VERSION : 0.1
   VAR_INPUT
      OFF_SQ : Bool := false;   // Turn sequence off
      INIT_SQ : Bool := false;   // Set sequence to initial state
      ACK_EF : Bool := false;   // Acknowledge all errors and faults
   END_VAR
   VAR_OUTPUT
      S_NO : Int := 0;   // Step number
      S_MORE : Bool := false;   // More steps are available and can be shown in S_NO
      S_ACTIVE : Bool := false;   // Step indicated in S_NO is active
      ERR_FLT : Bool := false;   // Interlock or supervision group error
      AUTO_ON : Bool := false;   // Automatic mode is active
   END_VAR
   VAR
      STATE : Int;   // Step number
      Unit : Struct
         START : Bool;   // Sequence Start
         INITIALIZATION : Bool;   // Sequence initialization
         ABORTING : Bool;   // Sequence about
         WAIT : Bool;   // Wating for Permissive read only
         COMPLETE : Bool;   // Sequence done
         "TURN ON" : Bool;   // Operator turn on retail equiment Button
         "TURN OFF" : Bool;   // Operator turn off retail equiment Button
         DONE : Bool;   // Operator Material is Being remove Button
         LV : Bool;
         PM : Bool;
         OverFlowCheck : Struct   // Check the Centrifuge is not over Material
            Enable : Bool;
            Wait_over : Bool;
            wait_pmp : Bool;
         END_STRUCT;
         TURBIDITY : Struct
            Enable : Bool;
            Wait : Bool;
         END_STRUCT;
         "WET CAKE_DRAIN" : Bool;
         Flow_SP : Real := 5.0;   // L/Min Flow Setpoint for FV-3011
         "TIMER" : Struct
            BucketTimer : IEC_TIMER;
            "WET-CAKE" : IEC_TIMER;
         END_STRUCT;
         "TIME" : Struct
            "WET-CAKE" : Time := T#10M;
            CountDown : Struct
               "WET-CAKE" : Time;
            END_STRUCT;
         END_STRUCT;
      END_STRUCT;
      HMI_INFO : Array[0..11] of UInt;
      IF_PAR : G7_IfParPlus_V6;
      RT_DATA : G7_RTDataPlus_V6;   // Internal data area
      Abort : G7_TransitionPlus_V6;   // Transition structure
      InitializeR : G7_TransitionPlus_V6;   // Transition structure
      CentfgP : G7_TransitionPlus_V6;   // Transition structure
      Re : G7_TransitionPlus_V6;   // Transition structure
      Centrifuge : G7_TransitionPlus_V6;   // Transition structure
      Wash : G7_TransitionPlus_V6;   // Transition structure
      Std : G7_TransitionPlus_V6;   // Transition structure
      StT : G7_TransitionPlus_V6;   // Transition structure
      MotorOn : G7_TransitionPlus_V6;   // Transition structure
      ROpnd : G7_TransitionPlus_V6;   // Transition structure
      AutoFlw : G7_TransitionPlus_V6;   // Transition structure
      TOT_Dn : G7_TransitionPlus_V6;   // Transition structure
      TransfDn : G7_TransitionPlus_V6;   // Transition structure
      TnkIdle : G7_TransitionPlus_V6;   // Transition structure
      WaterDn : G7_TransitionPlus_V6;   // Transition structure
      WtPmOff : G7_TransitionPlus_V6;   // Transition structure
      BcketTDn : G7_TransitionPlus_V6;   // Transition structure
      PmpsOff : G7_TransitionPlus_V6;   // Transition structure
      CntrfgOff : G7_TransitionPlus_V6;   // Transition structure
      CntrfgEnd : G7_TransitionPlus_V6;   // Transition structure
      Init : G7_TransitionPlus_V6;   // Transition structure
      SAut : G7_TransitionPlus_V6;   // Transition structure
      SIn : G7_TransitionPlus_V6;   // Transition structure
      Initd : G7_TransitionPlus_V6;   // Transition structure
      Trans145 : G7_TransitionPlus_V6;   // Transition structure
      Ab : G7_TransitionPlus_V6;   // Transition structure
      AbortOn : G7_TransitionPlus_V6;   // Transition structure
      AbortDn : G7_TransitionPlus_V6;   // Transition structure
      Idle : G7_StepPlus_V6;   // Step structure
      Ready : G7_StepPlus_V6;   // Step structure
      SelectSeq : G7_StepPlus_V6;   // Step structure
      Started : G7_StepPlus_V6;   // Step structure
      StartTank : G7_StepPlus_V6;   // Step structure
      "USER CentrOn" : G7_StepPlus_V6;   // Step structure
      OpenRoute : G7_StepPlus_V6;   // Step structure
      AutoFlowCtl : G7_StepPlus_V6;   // Step structure
      Transfering : G7_StepPlus_V6;   // Step structure
      Complete : G7_StepPlus_V6;   // Step structure
      ReleaseTank : G7_StepPlus_V6;   // Step structure
      "USER SlWash" : G7_StepPlus_V6;   // Step structure
      StopReqWater : G7_StepPlus_V6;   // Step structure
      Drying : G7_StepPlus_V6;   // Step structure
      DryingDone : G7_StepPlus_V6;   // Step structure
      "USER CentrOff" : G7_StepPlus_V6;   // Step structure
      End : G7_StepPlus_V6;   // Step structure
      Initialize : G7_StepPlus_V6;   // Step structure
      SetAuto : G7_StepPlus_V6;   // Step structure
      SetInitial : G7_StepPlus_V6;   // Step structure
      "2ndReset" : G7_StepPlus_V6;   // Step structure
      FeelerEngage : G7_StepPlus_V6;   // Step structure
      AbortStarting : G7_StepPlus_V6;   // Step structure
      Aborting : G7_StepPlus_V6;   // Step structure
      AbortDone : G7_StepPlus_V6;   // Step structure
      SINI : Array[0..4] of USInt;
      LSTT : Array[0..27] of USInt;
      ATAJ : Array[0..27] of USInt;
      ATAB : Array[0..27] of USInt;
      PSTT : Array[0..27] of USInt;
      NSTT : Array[0..27] of USInt;
      ASSJ : Array[0..24] of USInt;
      ASSB : Array[0..24] of USInt;
      PTTS : Array[0..24] of USInt;
      NTTS : Array[0..24] of USInt;
      SW_SQTS : Array[0..24] of USInt;
      SWITCH : Array[0..3] of USInt;
      TVX : Array[0..9] of USInt;
      TTX : Array[0..9] of USInt;
      TSX : Array[0..4] of USInt;
      S00X : Array[0..4] of USInt;
      SOFFX : Array[0..4] of USInt;
      SONX : Array[0..4] of USInt;
      SAX : Array[0..4] of USInt;
      SERRX : Array[0..25] of USInt;
      SMX : Array[0..25] of USInt;
      S0X : Array[0..25] of USInt;
      S1X : Array[0..25] of USInt;
      IL_ALARM_INST : Diag_Alarm;
      SUP_ALARM_INST : Diag_Alarm;
      STEP_TIME_ALARM_INST : Diag_Alarm;
      IEC_TIMER_INST : IEC_TIMER;
      TRANSACTION_FLAG : Bool := false;
   END_VAR
   // LSTT[8] := 255;
   // SINI[0] := 2;
   // LSTT[0] := 22;
   // NSTT[0] := 22;
   // PTTS[0] := 255;
   // TVX[0] := 16#1;
   // TTX[0] := 16#1;
   // TSX[0] := 16#1;
   // S00X[0] := 16#1;
   // SOFFX[0] := 16#1;
   // SONX[0] := 16#1;
   // SAX[0] := 16#1;
   // SERRX[0] := 16#1;
   // SMX[0] := 16#1;
   // S0X[0] := 16#1;
   // S1X[0] := 16#1;
   // LSTT[1] := 17;
   // LSTT[2] := 255;
   // LSTT[3] := 255;
   // LSTT[4] := 3;
   // LSTT[5] := 255;
   // LSTT[6] := 255;
   // LSTT[7] := 255;
   // LSTT[9] := 255;
   // LSTT[13] := 255;
   // LSTT[10] := 255;
   // LSTT[11] := 255;
   // LSTT[12] := 255;
   // NSTT[8] := 6;
   // LSTT[14] := 255;
   // LSTT[15] := 255;
   // LSTT[16] := 255;
   // LSTT[17] := 255;
   // LSTT[18] := 255;
   // ATAJ[1] := 1;
   // ATAJ[2] := 2;
   // ATAJ[3] := 3;
   // ATAJ[4] := 4;
   // ATAJ[5] := 5;
   // ATAJ[6] := 6;
   // ATAJ[7] := 7;
   // ATAJ[8] := 8;
   // ATAJ[9] := 9;
   // ATAJ[10] := 10;
   // ATAJ[11] := 11;
   // ATAJ[12] := 12;
   // ATAJ[13] := 13;
   // ATAJ[14] := 14;
   // ATAJ[15] := 15;
   // ATAJ[16] := 16;
   // ATAJ[17] := 17;
   // ATAJ[18] := 18;
   // ATAJ[19] := 19;
   // ATAB[1] := 2;
   // ATAB[17] := 17;
   // ATAB[3] := 3;
   // ATAB[4] := 5;
   // ATAB[5] := 4;
   // ATAB[6] := 6;
   // ATAB[7] := 7;
   // ATAB[8] := 8;
   // ATAB[9] := 9;
   // ATAB[10] := 10;
   // ATAB[11] := 11;
   // ATAB[12] := 12;
   // ATAB[13] := 13;
   // ATAB[14] := 14;
   // ATAB[15] := 15;
   // ATAB[16] := 16;
   // ATAB[19] := 19;
   // ATAB[18] := 18;
   // PSTT[17] := 14;
   // PSTT[14] := 11;
   // PSTT[3] := 1;
   // PSTT[4] := 2;
   // PSTT[5] := 2;
   // PSTT[6] := 3;
   // PSTT[7] := 4;
   // PSTT[8] := 5;
   // PSTT[9] := 6;
   // PSTT[10] := 7;
   // PSTT[11] := 8;
   // PSTT[12] := 9;
   // PSTT[13] := 10;
   // PSTT[15] := 12;
   // PSTT[16] := 13;
   // PSTT[19] := 16;
   // PSTT[18] := 15;
   // PSTT[21] := 18;
   // NSTT[1] := 17;
   // NSTT[2] := 1;
   // NSTT[3] := 2;
   // NSTT[4] := 3;
   // NSTT[5] := 255;
   // NSTT[6] := 4;
   // NSTT[7] := 5;
   // NSTT[9] := 7;
   // NSTT[13] := 11;
   // NSTT[10] := 8;
   // NSTT[11] := 9;
   // NSTT[12] := 10;
   // NSTT[14] := 12;
   // NSTT[15] := 13;
   // NSTT[16] := 14;
   // NSTT[17] := 15;
   // NSTT[18] := 16;
   // ASSJ[1] := 1;
   // ASSJ[2] := 2;
   // ASSJ[3] := 3;
   // ASSJ[4] := 4;
   // ASSJ[5] := 5;
   // ASSJ[6] := 6;
   // ASSJ[7] := 7;
   // ASSJ[8] := 8;
   // ASSJ[9] := 9;
   // ASSJ[10] := 10;
   // ASSJ[11] := 11;
   // ASSJ[12] := 12;
   // ASSJ[13] := 13;
   // ASSJ[14] := 14;
   // ASSJ[15] := 15;
   // ASSJ[16] := 16;
   // ASSB[1] := 1;
   // ASSB[2] := 2;
   // ASSB[3] := 3;
   // ASSB[4] := 4;
   // ASSB[5] := 5;
   // ASSB[6] := 6;
   // ASSB[7] := 7;
   // ASSB[8] := 8;
   // ASSB[9] := 9;
   // ASSB[10] := 10;
   // ASSB[11] := 11;
   // ASSB[12] := 12;
   // ASSB[13] := 13;
   // ASSB[14] := 14;
   // ASSB[15] := 15;
   // ASSB[16] := 16;
   // PTTS[2] := 3;
   // PTTS[3] := 255;
   // PTTS[4] := 6;
   // PTTS[5] := 7;
   // PTTS[6] := 8;
   // PTTS[7] := 9;
   // PTTS[8] := 10;
   // PTTS[9] := 11;
   // PTTS[10] := 12;
   // PTTS[11] := 13;
   // PTTS[12] := 14;
   // PTTS[13] := 15;
   // PTTS[14] := 16;
   // PTTS[15] := 17;
   // PTTS[16] := 18;
   // NTTS[1] := 3;
   // NTTS[2] := 4;
   // NTTS[3] := 6;
   // NTTS[4] := 7;
   // NTTS[5] := 8;
   // NTTS[6] := 9;
   // NTTS[7] := 10;
   // NTTS[8] := 11;
   // NTTS[9] := 12;
   // NTTS[10] := 13;
   // NTTS[11] := 14;
   // NTTS[12] := 15;
   // NTTS[13] := 16;
   // NTTS[14] := 17;
   // NTTS[15] := 18;
   // NTTS[16] := 19;
   // SW_SQTS[6] := 2;
   // SW_SQTS[7] := 2;
   // SW_SQTS[8] := 2;
   // SW_SQTS[9] := 2;
   // SW_SQTS[10] := 2;
   // SW_SQTS[11] := 2;
   // SW_SQTS[12] := 2;
   // SW_SQTS[13] := 2;
   // SW_SQTS[14] := 2;
   // SW_SQTS[15] := 2;
   // SW_SQTS[16] := 2;
   // NTTS[23] := 26;
   // NTTS[22] := 25;
   // NTTS[21] := 24;
   // NTTS[20] := 23;
   // NTTS[19] := 22;
   // NTTS[18] := 21;
   // NTTS[17] := 20;
   // PTTS[23] := 25;
   // PTTS[22] := 255;
   // PTTS[21] := 23;
   // PTTS[20] := 22;
   // PTTS[19] := 21;
   // PTTS[18] := 20;
   // PTTS[17] := 255;
   // ASSB[23] := 23;
   // ASSB[22] := 22;
   // ASSB[21] := 21;
   // ASSB[20] := 20;
   // ASSB[19] := 19;
   // ASSB[18] := 18;
   // ASSB[17] := 17;
   // ASSJ[23] := 23;
   // ASSJ[22] := 22;
   // ASSJ[21] := 21;
   // ASSJ[20] := 20;
   // ASSJ[19] := 19;
   // ASSJ[18] := 18;
   // ASSJ[17] := 17;
   // NSTT[23] := 21;
   // NSTT[25] := 23;
   // PSTT[26] := 23;
   // PSTT[25] := 22;
   // PSTT[24] := 21;
   // PSTT[23] := 20;
   // PSTT[22] := 19;
   // PSTT[20] := 17;
   // ATAB[26] := 26;
   // ATAB[25] := 25;
   // ATAB[24] := 24;
   // ATAB[23] := 23;
   // ATAB[22] := 22;
   // ATAB[21] := 21;
   // ATAB[20] := 20;
   // ATAJ[26] := 26;
   // ATAJ[25] := 25;
   // ATAJ[24] := 24;
   // ATAJ[23] := 23;
   // ATAJ[22] := 22;
   // ATAJ[21] := 21;
   // ATAJ[20] := 20;
   // LSTT[23] := 255;
   // LSTT[25] := 255;
   // SW_SQTS[17] := 3;
   // SW_SQTS[18] := 3;
   // SW_SQTS[19] := 3;
   // SW_SQTS[20] := 3;
   // SW_SQTS[21] := 3;
   // SW_SQTS[22] := 4;
   // SW_SQTS[23] := 4;
   // SINI[2] := 255;
   // SINI[3] := 255;
   // LSTT[21] := 255;
   // NSTT[21] := 19;
   // SW_SQTS[2] := 1;
   // SW_SQTS[3] := 2;
   // SW_SQTS[4] := 2;
   // SW_SQTS[5] := 2;
   // Unit."TIMER".BucketTimer.PT := T#10S;
   // LSTT[24] := 1;
   // LSTT[22] := 255;
   // NSTT[22] := 20;
   // NSTT[24] := 1;
   // Unit."TIMER"."WET-CAKE".PT := T#10M;
   // SINI[4] := 255;
   // LSTT[20] := 255;
   // NSTT[20] := 18;
   // PTTS[1] := 2;
   // SWITCH[1] := 239;
   // SWITCH[0] := 156;
   // SWITCH[2] := 251;
   // ATAB[0] := 1;
   // SW_SQTS[1] := 1;
   // LSTT[26] := 255;
   // ATAJ[27] := 27;
   // ATAB[27] := 27;
   // PSTT[27] := 24;
   // NSTT[26] := 24;
   // ASSJ[24] := 24;
   // ASSB[24] := 24;
   // PTTS[24] := 26;
   // NTTS[24] := 27;
   // SW_SQTS[24] := 4;
BEGIN
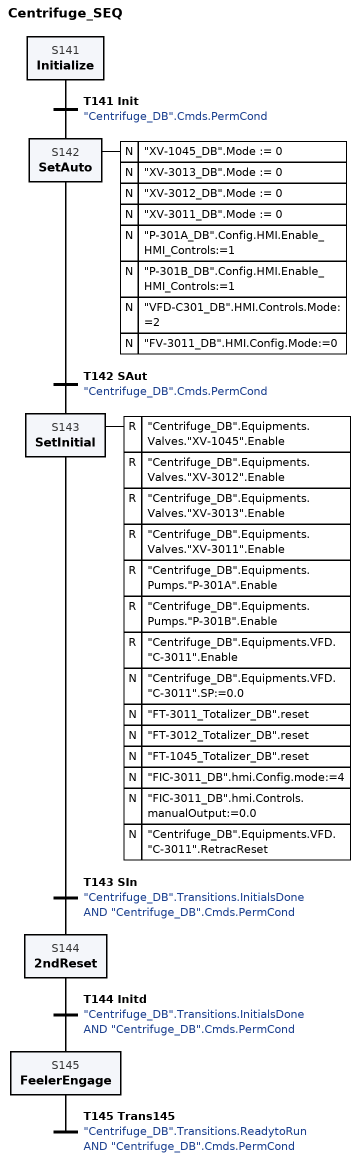
   // permanent pre-instructions
   NETWORK 1
      "Centrifuge_Signals_FROM_T-103"();
      "Centrifuge_Signals_FROM_T-104"();
      "Centrifuge_SEQ_FC"();
      "Centrifuge_Transitions_FC"();

   // sequencer 1
   STEP "2ndReset":   // S144, max time T#10S, warning time T#7S
      // Initialize T-101 Batch sequence
   END_STEP
   TRANSITION Initd FROM "2ndReset" TO FeelerEngage   // T144
      := "Centrifuge_DB".Transitions.InitialsDone AND "Centrifuge_DB".Cmds.PermCond;
   END_TRANSITION
   STEP Initialize:   // S141, max time T#10S, warning time T#7S
      // Initialize T-101 Batch sequence
   END_STEP
   TRANSITION Init FROM Initialize TO SetAuto   // T141: CLOSED: XV-1041
      := "Centrifuge_DB".Cmds.PermCond;
   END_TRANSITION
   STEP SetInitial:   // S143, max time T#10S, warning time T#7S
      // Initialize T-101 Batch sequence
              R    "Centrifuge_DB".Equipments.Valves."XV-1045".Enable
              R    "Centrifuge_DB".Equipments.Valves."XV-3012".Enable
              R    "Centrifuge_DB".Equipments.Valves."XV-3013".Enable
              R    "Centrifuge_DB".Equipments.Valves."XV-3011".Enable
              R    "Centrifuge_DB".Equipments.Pumps."P-301A".Enable
              R    "Centrifuge_DB".Equipments.Pumps."P-301B".Enable
              R    "Centrifuge_DB".Equipments.VFD."C-3011".Enable
              N    "Centrifuge_DB".Equipments.VFD."C-3011".SP:=0.0
              N    "FT-3011_Totalizer_DB".reset
              N    "FT-3012_Totalizer_DB".reset
              N    "FT-1045_Totalizer_DB".reset
              N    "FIC-3011_DB".hmi.Config.mode:=4
              N    "FIC-3011_DB".hmi.Controls.manualOutput:=0.0
              N    "Centrifuge_DB".Equipments.VFD."C-3011".RetracReset
   END_STEP
   TRANSITION SIn FROM SetInitial TO "2ndReset"   // T143: CLOSED: XV-1013
      := "Centrifuge_DB".Transitions.InitialsDone AND "Centrifuge_DB".Cmds.PermCond;
   END_TRANSITION
   STEP SetAuto:   // S142, max time T#10S, warning time T#7S
              N    "XV-1045_DB".Mode := 0
              N    "XV-3013_DB".Mode := 0
              N    "XV-3012_DB".Mode := 0
              N    "XV-3011_DB".Mode := 0
              N    "P-301A_DB".Config.HMI.Enable_HMI_Controls:=1
              N    "P-301B_DB".Config.HMI.Enable_HMI_Controls:=1
              N    "VFD-C301_DB".HMI.Controls.Mode:=2
              N    "FV-3011_DB".HMI.Config.Mode:=0
   END_STEP
   TRANSITION SAut FROM SetAuto TO SetInitial   // T142
      := "Centrifuge_DB".Cmds.PermCond;
   END_TRANSITION
   STEP FeelerEngage:   // S145, max time T#10S, warning time T#7S
   END_STEP
   TRANSITION Trans145 FROM FeelerEngage TO ?   // T145
      := "Centrifuge_DB".Transitions.ReadytoRun AND "Centrifuge_DB".Cmds.PermCond;
   END_TRANSITION

   // permanent post-instructions
   NETWORK 1
      "Centrifuge_FC_Outputs"();
END_FUNCTION_BLOCK

FUNCTION "Centrifuge_SEQ_FC_old" : Void   // FC75, LAD
{ S7_Optimized_Access := 'TRUE' }
VERSION : 0.1
   VAR_TEMP   // added for the SCL form of the ladder/FBD networks
      _w1 : Bool;
      _w2 : Bool;
   END_VAR
BEGIN

REGION Network 2: Abort
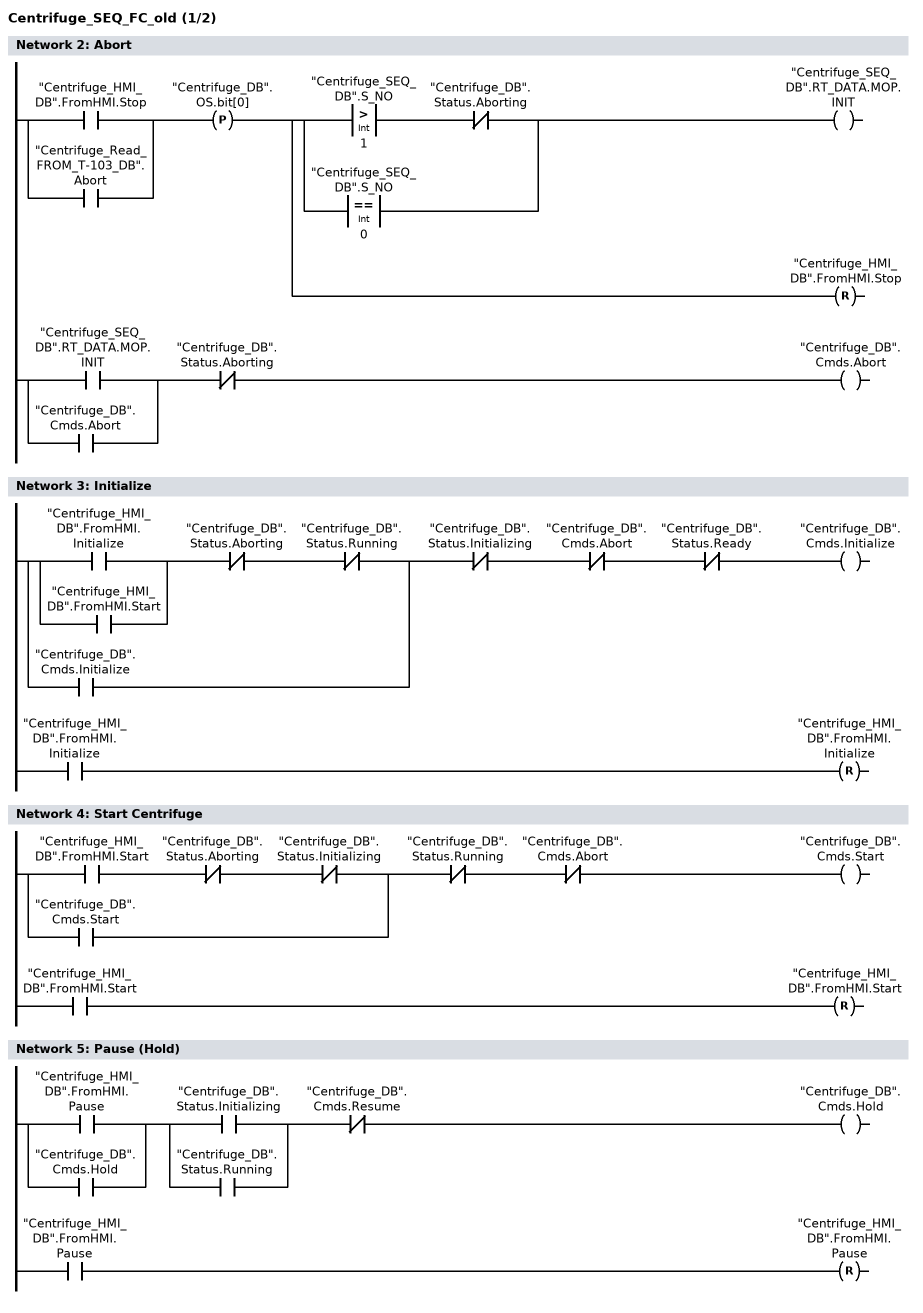
   RUNG wire#powerrail
      Contact( "Centrifuge_HMI_DB".FromHMI.Stop )
      wire#w1
      P_Trig( "Centrifuge_DB".OS.bit[0] )
      wire#w2
      { S7_Templates := "SrcType := Int" } GT_Contact(in1 := "Centrifuge_SEQ_DB".S_NO, in2 := 1)
      I_Contact( "Centrifuge_DB".Status.Aborting )
      wire#w3
      Coil( "Centrifuge_SEQ_DB".RT_DATA.MOP.INIT )
   END_RUNG
   RUNG wire#powerrail
      Contact( "Centrifuge_Read_FROM_T-103_DB".Abort )
   END_RUNG wire#w1
   RUNG wire#w2
      { S7_Templates := "SrcType := Int" } EQ_Contact(in1 := "Centrifuge_SEQ_DB".S_NO, in2 := 0)
   END_RUNG wire#w3
   RUNG wire#w2
      R_Coil( "Centrifuge_HMI_DB".FromHMI.Stop )
   END_RUNG
   RUNG wire#powerrail
      Contact( "Centrifuge_SEQ_DB".RT_DATA.MOP.INIT )
      wire#w4
      I_Contact( "Centrifuge_DB".Status.Aborting )
      Coil( "Centrifuge_DB".Cmds.Abort )
   END_RUNG
   RUNG wire#powerrail
      Contact( "Centrifuge_DB".Cmds.Abort )
   END_RUNG wire#w4
   // the same network as SCL:
   #_w1 := "Centrifuge_HMI_DB".FromHMI.Stop OR "Centrifuge_Read_FROM_T-103_DB".Abort;
   #_w2 := #_w1 AND NOT "Centrifuge_DB".OS.bit[0];   // rising edge
   "Centrifuge_DB".OS.bit[0] := #_w1;
   "Centrifuge_SEQ_DB".RT_DATA.MOP.INIT := #_w2 AND ((("Centrifuge_SEQ_DB".S_NO > 1) AND NOT "Centrifuge_DB".Status.Aborting) OR ("Centrifuge_SEQ_DB".S_NO = 0));
   IF #_w2 THEN "Centrifuge_HMI_DB".FromHMI.Stop := FALSE; END_IF;
   "Centrifuge_DB".Cmds.Abort := ("Centrifuge_SEQ_DB".RT_DATA.MOP.INIT OR "Centrifuge_DB".Cmds.Abort) AND NOT "Centrifuge_DB".Status.Aborting;
END_REGION

REGION Network 3: Initialize
   RUNG wire#powerrail
      Contact( "Centrifuge_HMI_DB".FromHMI.Initialize )
      wire#w1
      I_Contact( "Centrifuge_DB".Status.Aborting )
      I_Contact( "Centrifuge_DB".Status.Running )
      wire#w2
      I_Contact( "Centrifuge_DB".Status.Initializing )
      I_Contact( "Centrifuge_DB".Cmds.Abort )
      I_Contact( "Centrifuge_DB".Status.Ready )
      Coil( "Centrifuge_DB".Cmds.Initialize )
   END_RUNG
   RUNG wire#powerrail
      Contact( "Centrifuge_HMI_DB".FromHMI.Start )
   END_RUNG wire#w1
   RUNG wire#powerrail
      Contact( "Centrifuge_DB".Cmds.Initialize )
   END_RUNG wire#w2
   RUNG wire#powerrail
      Contact( "Centrifuge_HMI_DB".FromHMI.Initialize )
      R_Coil( "Centrifuge_HMI_DB".FromHMI.Initialize )
   END_RUNG
   // the same network as SCL:
   "Centrifuge_DB".Cmds.Initialize := ((("Centrifuge_HMI_DB".FromHMI.Initialize OR "Centrifuge_HMI_DB".FromHMI.Start) AND NOT "Centrifuge_DB".Status.Aborting AND NOT "Centrifuge_DB".Status.Running) OR "Centrifuge_DB".Cmds.Initialize) AND NOT "Centrifuge_DB".Status.Initializing AND NOT "Centrifuge_DB".Cmds.Abort AND NOT "Centrifuge_DB".Status.Ready;
   IF "Centrifuge_HMI_DB".FromHMI.Initialize THEN "Centrifuge_HMI_DB".FromHMI.Initialize := FALSE; END_IF;
END_REGION

REGION Network 4: Start Centrifuge
   RUNG wire#powerrail
      Contact( "Centrifuge_HMI_DB".FromHMI.Start )
      I_Contact( "Centrifuge_DB".Status.Aborting )
      I_Contact( "Centrifuge_DB".Status.Initializing )
      wire#w1
      I_Contact( "Centrifuge_DB".Status.Running )
      I_Contact( "Centrifuge_DB".Cmds.Abort )
      Coil( "Centrifuge_DB".Cmds.Start )
   END_RUNG
   RUNG wire#powerrail
      Contact( "Centrifuge_DB".Cmds.Start )
   END_RUNG wire#w1
   RUNG wire#powerrail
      Contact( "Centrifuge_HMI_DB".FromHMI.Start )
      R_Coil( "Centrifuge_HMI_DB".FromHMI.Start )
   END_RUNG
   // the same network as SCL:
   "Centrifuge_DB".Cmds.Start := (("Centrifuge_HMI_DB".FromHMI.Start AND NOT "Centrifuge_DB".Status.Aborting AND NOT "Centrifuge_DB".Status.Initializing) OR "Centrifuge_DB".Cmds.Start) AND NOT "Centrifuge_DB".Status.Running AND NOT "Centrifuge_DB".Cmds.Abort;
   IF "Centrifuge_HMI_DB".FromHMI.Start THEN "Centrifuge_HMI_DB".FromHMI.Start := FALSE; END_IF;
END_REGION

REGION Network 5: Pause (Hold)
   RUNG wire#powerrail
      Contact( "Centrifuge_HMI_DB".FromHMI.Pause )
      wire#w1
      Contact( "Centrifuge_DB".Status.Initializing )
      wire#w2
      I_Contact( "Centrifuge_DB".Cmds.Resume )
      Coil( "Centrifuge_DB".Cmds.Hold )
   END_RUNG
   RUNG wire#powerrail
      Contact( "Centrifuge_DB".Cmds.Hold )
   END_RUNG wire#w1
   RUNG wire#w1
      Contact( "Centrifuge_DB".Status.Running )
   END_RUNG wire#w2
   RUNG wire#powerrail
      Contact( "Centrifuge_HMI_DB".FromHMI.Pause )
      R_Coil( "Centrifuge_HMI_DB".FromHMI.Pause )
   END_RUNG
   // the same network as SCL:
   "Centrifuge_DB".Cmds.Hold := ("Centrifuge_HMI_DB".FromHMI.Pause OR "Centrifuge_DB".Cmds.Hold) AND ("Centrifuge_DB".Status.Initializing OR "Centrifuge_DB".Status.Running) AND NOT "Centrifuge_DB".Cmds.Resume;
   IF "Centrifuge_HMI_DB".FromHMI.Pause THEN "Centrifuge_HMI_DB".FromHMI.Pause := FALSE; END_IF;
END_REGION

REGION Network 6: Restart From Pause (Hold)
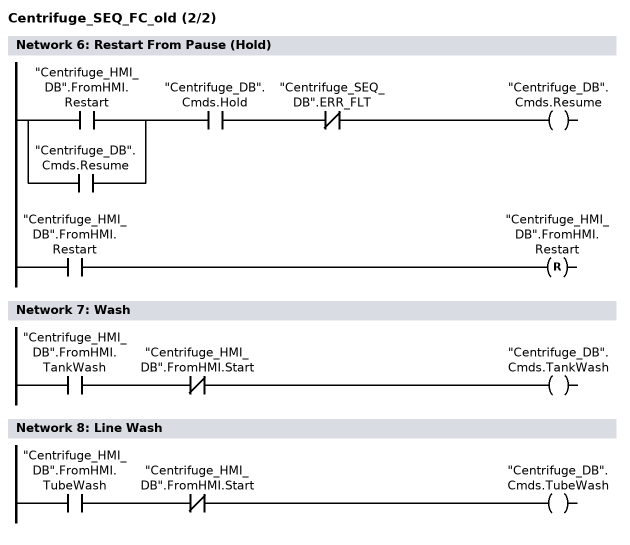
   RUNG wire#powerrail
      Contact( "Centrifuge_HMI_DB".FromHMI.Restart )
      wire#w1
      Contact( "Centrifuge_DB".Cmds.Hold )
      I_Contact( "Centrifuge_SEQ_DB".ERR_FLT )
      Coil( "Centrifuge_DB".Cmds.Resume )
   END_RUNG
   RUNG wire#powerrail
      Contact( "Centrifuge_DB".Cmds.Resume )
   END_RUNG wire#w1
   RUNG wire#powerrail
      Contact( "Centrifuge_HMI_DB".FromHMI.Restart )
      R_Coil( "Centrifuge_HMI_DB".FromHMI.Restart )
   END_RUNG
   // the same network as SCL:
   "Centrifuge_DB".Cmds.Resume := ("Centrifuge_HMI_DB".FromHMI.Restart OR "Centrifuge_DB".Cmds.Resume) AND "Centrifuge_DB".Cmds.Hold AND NOT "Centrifuge_SEQ_DB".ERR_FLT;
   IF "Centrifuge_HMI_DB".FromHMI.Restart THEN "Centrifuge_HMI_DB".FromHMI.Restart := FALSE; END_IF;
END_REGION

REGION Network 7: Wash
   RUNG wire#powerrail
      Contact( "Centrifuge_HMI_DB".FromHMI.TankWash )
      I_Contact( "Centrifuge_HMI_DB".FromHMI.Start )
      Coil( "Centrifuge_DB".Cmds.TankWash )
   END_RUNG
   // the same network as SCL:
   "Centrifuge_DB".Cmds.TankWash := "Centrifuge_HMI_DB".FromHMI.TankWash AND NOT "Centrifuge_HMI_DB".FromHMI.Start;
END_REGION

REGION Network 8: Line Wash
   RUNG wire#powerrail
      Contact( "Centrifuge_HMI_DB".FromHMI.TubeWash )
      I_Contact( "Centrifuge_HMI_DB".FromHMI.Start )
      Coil( "Centrifuge_DB".Cmds.TubeWash )
   END_RUNG
   // the same network as SCL:
   "Centrifuge_DB".Cmds.TubeWash := "Centrifuge_HMI_DB".FromHMI.TubeWash AND NOT "Centrifuge_HMI_DB".FromHMI.Start;
END_REGION

REGION Network 9 (SCL): Sequence Status
   IF "Centrifuge_SEQ_DB".S_NO= 1 THEN
       "Centrifuge_DB".Status.Status := 1; //Idle
   ELSIF "Centrifuge_SEQ_DB".S_NO > 1 AND "Centrifuge_SEQ_DB".S_NO < 150 AND NOT "Centrifuge_SEQ_DB".ERR_FLT THEN
       "Centrifuge_DB".Status.Status := 2; //Running
   ELSIF "Centrifuge_SEQ_DB".S_NO >= 151 AND "Centrifuge_SEQ_DB".S_NO <= 160 AND NOT "Centrifuge_SEQ_DB".ERR_FLT THEN
       "Centrifuge_DB".Status.Status := 3; // Stopping
   ELSIF ("Centrifuge_SEQ_DB".ERR_FLT OR "Centrifuge_DB".Cmds.Hold)  AND "Centrifuge_DB".Status.Status =2 THEN
       "Centrifuge_DB".Status.Status := 4; //Held
   ELSIF ("Centrifuge_SEQ_DB".ERR_FLT OR "Centrifuge_DB".Cmds.Hold) AND  "Centrifuge_DB".Status.Status =2 AND "Centrifuge_Aux_DB"."Bool".TOff  THEN
       "Centrifuge_DB".Status.Status := 5; // Holding
   ELSE
       "Centrifuge_DB".Status.Status := 6; //Unknown
   END_IF;

   //Enable/Disable HMI Start/Stop Button
   "Centrifuge_HMI_DB".ToHMI.EnStopButton := ("Centrifuge_DB".Status.Status > 1) OR "Centrifuge_DB".Status.Step = 0; //Enable HMI Stop Button
   "Centrifuge_HMI_DB".ToHMI.EnStartButton := "Centrifuge_DB".Status.Status = 1;   //Enable Start Button
   "Centrifuge_HMI_DB".ToHMI.EnPauseButton := "Centrifuge_DB".Status.Status = 2 AND NOT "Centrifuge_DB".Cmds.Hold; //Enable Pause Button
   "Centrifuge_HMI_DB".ToHMI.EnRestartButton := "Centrifuge_DB".Status.Status = 2 AND "Centrifuge_DB".Cmds.Hold; //Enable Restart Button
END_REGION

REGION Network 10 (SCL): Sequence Step
   "Centrifuge_DB".Status.Step := "Centrifuge_SEQ_DB".S_NO;
END_REGION

REGION Network 11 (SCL): Sequence state (Procedure running)
   IF "Centrifuge_SEQ_DB".S_NO = 3 OR "Centrifuge_SEQ_DB".S_NO = 4 THEN
       "Centrifuge_DB".Status.State := 1; //Ready
   ELSIF "Centrifuge_SEQ_DB".S_NO >= 21 AND "Centrifuge_SEQ_DB".S_NO <= 60 THEN
       "Centrifuge_DB".Status.State := 2; //Mixing 
   ELSIF "Centrifuge_SEQ_DB".S_NO >= 61 AND "Centrifuge_SEQ_DB".S_NO <= 80 THEN
       "Centrifuge_DB".Status.State := 3; //Pouring
   ELSIF "Centrifuge_SEQ_DB".S_NO >= 141 AND "Centrifuge_SEQ_DB".S_NO <= 150 THEN
       "Centrifuge_DB".Status.State := 4; //Initializing
   ELSIF "Centrifuge_SEQ_DB".S_NO >= 151 AND "Centrifuge_SEQ_DB".S_NO <= 160 THEN
       "Centrifuge_DB".Status.State := 5; //Aborting
   ELSE
       "Centrifuge_DB".Status.State := 0;
   END_IF;
END_REGION

REGION Network 12: Sequence State
END_REGION
END_FUNCTION

FUNCTION "Centrifuge_FC_Outputs" : Void   // FC84, SCL
{ S7_Optimized_Access := 'TRUE' }
VERSION : 0.1
   VAR_TEMP
      Pump_A : Struct
         Cond_01 : Bool;   // Condition 01
         Cond_02 : Bool;
         Cond_03 : Bool;
         Cond_04 : Bool;
      END_STRUCT;
      Pump_B : Struct
         Cond_01 : Bool;   // Condition 01
         Cond_02 : Bool;   // Condition 02
         Cond_03 : Bool;
         Cond_04 : Bool;
         Cond_05 : Bool;
      END_STRUCT;
      Motor : Struct
         Cond_01 : Bool;   // Condition 01
         Cond_02 : Bool;   // Condition 02
      END_STRUCT;
      XV : Struct
         "1045" : Bool;
         "3011" : Bool;
         "3012" : Bool;
         "3013" : Bool;
      END_STRUCT;
      "FV-3011" : Struct
         On : Bool;
         Cond_1 : Bool;
      END_STRUCT;
   END_VAR
BEGIN
   //****** Equipmens Activation*******
   //
   //**************************************************************
   //

   //IF "AlwaysFALSE"  AND  ("Centrifuge_DB".Status.Status <> 1) THEN

       //***********************************************Water Inlet Valve**********************************************************************
       IF "XV-1045_DB".Mode = 0 THEN
           "Centrifuge_DB".Equipments.Valves."XV-1045".CmdOn := "Centrifuge_DB".Equipments.Valves."XV-1045".Enable 
           AND "ZT-C301_DB".SAI>"CentrifugeSpeed" AND NOT "Centrifuge_DB".Cmds.Hold;
           //Delay Off To avoid Overpressure the Lines
           #XV."1045" := "Centrifuge_DB".Equipments.Valves."XV-1045".CmdOn;
           "Centrifuge_Aux_DB".Timer."XV-1045".TOF(IN := #XV."1045",
                                                   PT := "Centrifuge_Aux_DB".Constants.CmdDelay);
           //Command to the Valve
           IF "Centrifuge_Aux_DB".Timer."XV-1045".Q THEN
               "XV-1045_DB".CMD := 2;
           ELSE
               "XV-1045_DB".CMD := 1;
           END_IF;
           "Centrifuge_DB".Equipments.Valves."XV-1045".TurningOff := NOT "Centrifuge_DB".Equipments.Valves."XV-1045".CmdOn AND "Centrifuge_Aux_DB".Timer."XV-1045".Q;
       END_IF;
       //***********************************************Inlet Valve**********************************************************************
       IF "XV-3011_DB".Mode = 0 THEN
           "Centrifuge_DB".Equipments.Valves."XV-3011".CmdOn := "Centrifuge_DB".Equipments.Valves."XV-3011".Enable
           AND NOT "Centrifuge_Aux_DB"."Bool".Centrifuge.Status.FeelerRetracted  AND NOT "Centrifuge_DB".Cmds.Hold;
           //Delay Off To avoid Overpressure the Lines
           #XV."3011" := "Centrifuge_DB".Equipments.Valves."XV-3011".CmdOn;
           "Centrifuge_Aux_DB".Timer."XV-3011".TOF(IN := #XV."3011",
           PT := "Centrifuge_Aux_DB".Constants.CmdDelay);
           IF "Centrifuge_Aux_DB".Timer."XV-3011".Q THEN
               "XV-3011_DB".CMD := 2;
           ELSE
               "XV-3011_DB".CMD := 1;
           END_IF;
           "Centrifuge_DB".Equipments.Valves."XV-3011".TurningOff := NOT "Centrifuge_DB".Equipments.Valves."XV-3011".CmdOn AND "Centrifuge_Aux_DB".Timer."XV-3011".Q;
       END_IF;
       //***********************************************Return Valve**********************************************************************
       IF "XV-3012_DB".Mode = 0 THEN
           "Centrifuge_DB".Equipments.Valves."XV-3012".CmdOn := "Centrifuge_DB".Equipments.Valves."XV-3012".Enable AND NOT "Centrifuge_DB".Cmds.Hold;
           //Delay Off To avoid Overpressure the Lines
           #XV."3012" := "Centrifuge_DB".Equipments.Valves."XV-3012".CmdOn;
           "Centrifuge_Aux_DB".Timer."XV-3012".TOF(IN := #XV."3012",
                                                   PT := "Centrifuge_Aux_DB".Constants.CmdDelay);
           //Command to the Valve
           IF "Centrifuge_Aux_DB".Timer."XV-3012".Q THEN
               "XV-3012_DB".CMD := 2;
           ELSE
               "XV-3012_DB".CMD := 1;
           END_IF;
           "Centrifuge_DB".Equipments.Valves."XV-3012".TurningOff := NOT "Centrifuge_DB".Equipments.Valves."XV-3012".CmdOn AND "Centrifuge_Aux_DB".Timer."XV-3012".Q;
       END_IF;
       //***********************************************Outlet Valve**********************************************************************
       IF "XV-3013_DB".Mode = 0 THEN
           "Centrifuge_DB".Equipments.Valves."XV-3013".CmdOn := "Centrifuge_DB".Equipments.Valves."XV-3013".Enable AND NOT "Centrifuge_DB".Cmds.Hold;
           //Delay Off To avoid Overpressure the Lines
           #XV."3013" := "Centrifuge_DB".Equipments.Valves."XV-3013".CmdOn;
           "Centrifuge_Aux_DB".Timer."XV-3013".TOF(IN := #XV."3013",
                                                   PT := "Centrifuge_Aux_DB".Constants.CmdDelay);
           //Command to the Valve
           IF "Centrifuge_Aux_DB".Timer."XV-3013".Q THEN
               "XV-3013_DB".CMD := 2;
           ELSE
               "XV-3013_DB".CMD := 1;
           END_IF;
           "Centrifuge_DB".Equipments.Valves."XV-3013".TurningOff := NOT "Centrifuge_DB".Equipments.Valves."XV-3013".CmdOn AND "Centrifuge_Aux_DB".Timer."XV-3013".Q;
       END_IF;

       //***********************************************FIC-3011 Controller (Centrifuge inlet flow)********************************************************************
       IF "FV-3011_DB".HMI.Config.Mode = 0 THEN
           #"FV-3011".Cond_1 := "Centrifuge_DB".Equipments.Valves."FV-3011".Enable AND "XV-3011_DB".OS;
           "Centrifuge_DB".Equipments.Valves."FV-3011".CmdOn := #"FV-3011".Cond_1 AND NOT "Centrifuge_DB".Cmds.Hold AND NOT "Centrifuge_DB".Status.Aborting;
           //Delay Off To avoid Overpressure the Lines
           #"FV-3011".On := "Centrifuge_DB".Equipments.Valves."FV-3011".CmdOn;
           "Centrifuge_Aux_DB".Timer."FV-3011".TOF(IN := #"FV-3011".On,
                                                   PT := "Centrifuge_Aux_DB".Constants.CmdDelay);
           IF "Centrifuge_Aux_DB".Timer."FV-3011".Q THEN
               "FIC-3011_DB".enableManualMode := False;
               "FIC-3011_DB".enableRemoteSetpoint := False;
               "FIC-3011_DB".hmi.Controls.manualEnable := False;
               "FIC-3011_DB".hmi.Config.mode := 3;
           END_IF;     // ELSE
             //  "FIC-3011_DB".enableManualMode := True;
             //  "FIC-3011_DB".enableRemoteSetpoint := False;
             //  "FIC-3011_DB".hmi.Controls.manualEnable := True;
             //  "FIC-3011_DB".hmi.Config.mode := 4;
            //   "FIC-3011_DB".hmi.Controls.manualOutput := 0;
         //  END_IF;
           "Centrifuge_DB".Equipments.Valves."FV-3011".TurningOff := NOT "Centrifuge_DB".Equipments.Valves."FV-3011".CmdOn AND "Centrifuge_Aux_DB".Timer."FV-3011".Q;
       END_IF;
       // ***********************************************Pump A**********************************************************************
       // Condition to CmdOn "On Command" 
       IF "P-301A_DB".Config.HMI.Enable_HMI_Controls = 1 THEN
           #Pump_A.Cond_01 := "Centrifuge_DB".Equipments.Pumps."P-301A".Enable AND ("Centrifuge_DB".PmpSel."P-301AB" = 1 OR "Centrifuge_DB".PmpSel."P-301AB" = 3);
           #Pump_A.Cond_02 :=  "XV-3013_DB".OS OR "XV-3012_DB".OS; //Outlet Valve Open. 
           #Pump_A.Cond_03 := #Pump_A.Cond_01 AND NOT "Centrifuge_DB".Cmds.Hold;
           "Centrifuge_DB".Equipments.Pumps."P-301A".CmdOn := #Pump_A.Cond_02 AND #Pump_A.Cond_03;
           //**********Commands to the Pumps
           IF "Centrifuge_DB".Equipments.Pumps."P-301A".CmdOn THEN
               "P-301A_DB".Stop_CMD := False;
               "P-301A_DB".Start_CMD := true;
               "P-301A_DB".ON := TRUE;
               "P-301A_DB".OFF := FALSE;
           ELSE
               "P-301A_DB".Stop_CMD := TRUE;
               "P-301A_DB".Start_CMD := FALSE;
               "P-301A_DB".ON := FALSE;
               "P-301A_DB".OFF := TRUE;
           END_IF;
       END_IF;
       // ***********************************************Pump B**********************************************************************
       // Condition to CmdOn "On Command" 
       IF "P-301B_DB".Config.HMI.Enable_HMI_Controls = 1 THEN
           #Pump_B.Cond_01 := "Centrifuge_DB".Equipments.Pumps."P-301B".Enable AND ("Centrifuge_DB".PmpSel."P-301AB" = 2 OR "Centrifuge_DB".PmpSel."P-301AB" = 3);
           #Pump_B.Cond_02 := "XV-3013_DB".OS OR "XV-3012_DB".OS; //Outlet Valve Open. 
           #Pump_B.Cond_03 := #Pump_B.Cond_01 AND NOT "Centrifuge_DB".Cmds.Hold;
           "Centrifuge_DB".Equipments.Pumps."P-301B".CmdOn := #Pump_B.Cond_02 AND #Pump_B.Cond_03;
           //**********Commands to the Pumps
           IF "Centrifuge_DB".Equipments.Pumps."P-301B".CmdOn THEN
               "P-301B_DB".Stop_CMD := False;
               "P-301B_DB".Start_CMD := true;
               "P-301B_DB".ON := TRUE;
               "P-301B_DB".OFF := FALSE;
           ELSE
               "P-301B_DB".Stop_CMD := TRUE;
               "P-301B_DB".Start_CMD := FALSE;
               "P-301B_DB".ON := FALSE;
               "P-301B_DB".OFF := TRUE;
           END_IF;
       END_IF;
       //***********************************************Motor**********************************************************************
       IF "VFD-C301_DB".HMI.Controls.Mode = 2 THEN
           #Motor.Cond_01 := "Centrifuge_DB".Equipments.VFD."C-3011".Enable;
           #Motor.Cond_02 := "AlwaysTRUE";
           "Centrifuge_DB".Equipments.VFD."C-3011".Start := #Motor.Cond_01 AND #Motor.Cond_02 AND NOT "Centrifuge_DB".Cmds.Hold;

           IF "Centrifuge_DB".Equipments.VFD."C-3011".Start THEN
               "VFD-C301_DB".PLCCommand := TRUE;
           ELSE
               "VFD-C301_DB".PLCCommand := FALSE;
           END_IF;
       END_IF;


      // END_IF;

       //*************************************************Transitions*************************************************
       "Centrifuge_DB".Transitions.WaterDone :="Centrifuge_DB".Status.Step = 30 AND "Centrifuge_Read_FROM_T-104_DB".PumpsOff AND "FT-1045_DB".SAI < 0.2;
       //*************************************************Interlocks to T-103*************************************************
       "Centrifuge_Write_TO_T-103_DB".RouteOpened := ("Centrifuge_DB".Status.Step = 24 OR "Centrifuge_DB".Status.Step = 25 OR "Centrifuge_DB".Status.Step = 26) AND "XV-3011_DB".OS AND ("FV-3011_DB".CMD > 80)
       AND ("XV-3013_DB".OS OR "XV-3012_DB".OS) AND "ZT-C301_DB".SAI>"CentrifugeSpeed";

       "Centrifuge_Write_TO_T-103_DB"."T-103_Empty" := "Centrifuge_DB".Status.Step = 27 AND "Centrifuge_DB".Transitions."T-103_Empty"
       AND NOT "Centrifuge_DB".Transitions.BasketFull;

       "Centrifuge_Write_TO_T-103_DB".BasketFull:= "Centrifuge_DB".Status.Step = 27 AND NOT "Centrifuge_DB".Transitions."T-103_Empty"
       AND "Centrifuge_DB".Transitions.BasketFull;

       "Centrifuge_Write_TO_T-103_DB".Release := "Centrifuge_DB".Status.Step = 28 AND NOT "Centrifuge_Read_FROM_T-103_DB".ReadyToTransfer;

       "Centrifuge_Write_TO_T-103_DB".FeelerRet := "Centrifuge_Aux_DB"."Bool".Centrifuge.Status.FeelerRetracted;